PopupScreen "Tank 2S Status" 885x425
   TrendView "Trend view_1" at 280,6 size 600x360
   TextField "Text field_4" at 20,134 size 86x22; Text 'Pressure:'
   IOField "I/O field_1" at 175,129 size 90x25; FormatPattern s999.9; Unit  mBar
      ProcessValue <- "20_TANKS_IP_DATA_RIO_02_FIRST_TANK_TANKS_PRESS"
   TextField "Text field_5" at 20,168 size 113x22; Text 'Water Level:'
   IOField "I/O field_2" at 175,163 size 90x25; FormatPattern 999.9; Unit  %
      ProcessValue <- "20_TANKS_IP_DATA_RIO_02_SECOND_TANK_BWT_LEVEL"
   TextField "Text field_6" at 20,202 size 137x22; Text 'MBG Flow Rate:'
   IOField "I/O field_3" at 175,197 size 90x25; FormatPattern 999.9; Unit  m³/hr
      ProcessValue <- "20_TANKS_IP_DATA_RIO_02_SECOND_TANK_MBG_FLOW"
   TextField "Text field_7" at 20,236 size 135x22; Text 'USD Flow Rate:'
   IOField "I/O field_4" at 175,231 size 90x25; FormatPattern 999.9; Unit  m³/hr
      ProcessValue <- "20_TANKS_IP_DATA_RIO_02_SECOND_TANK_USD_FLOW"
   TextField "Text field_8" at 20,270 size 140x22; Text 'Water pH Level:'
   IOField "I/O field_5" at 175,265 size 90x25; FormatPattern 99.9
      ProcessValue <- "20_TANKS_IP_DATA_RIO_02_SECOND_TANK_BWT_PH"
   TextField "Text field_9" at 20,304 size 143x22; Text 'Water DO Level:'
   IOField "I/O field_6" at 175,299 size 90x25; FormatPattern 99.99; Unit  mg/l
      ProcessValue <- "20_TANKS_IP_DATA_RIO_02_SECOND_TANK_BWT_DO"
   TextField "Text field_10" at 20,338 size 174x22; Text 'Water Temperature:'
   IOField "I/O field_7" at 190,333 size 75x25; FormatPattern 999.9; Unit  °C
      ProcessValue <- "20_TANKS_IP_DATA_RIO_02_SECOND_TANK_BWT_TEMP"
   Button "Button_4" at 550,375 size 150x40; TextOff 'Disable Tank'; Authorization "Operate"
      on Press: function_b14e0dd5("504_Tank Grouping_DB2020_TANK ACTIV 5", 0)
   Button "Button_1" at 50,5 size 220x35; TextOff 'Starboard Tank 2 (2S)'
      on Release: function_efd93a16("Tank 2S Status", 168, 315, -1, 0, 1)
   TextField "Text field_1" at 20,90 size 109x25; Text 'TIME LEFT:'
   GraphicView "Graphic view_1" at 20,46 size 245x32; Picture "Tank Manually Disabled"
   GraphicIOField "Graphic I/O field_1" at 20,46 size 245x32; PictureList "Tank Process Stage_II"
      Visibility <- "504_Tank Grouping_DB2020_GROUP of TANK 5"
      ProcessValue <- "2110_BTCS_CNTRL_DB_BTCS_STATE"
   Button "Button_2" at 4,5 size 45x35; TextOff 'Text'; PictureOff "Graphic_286"
      on Click: function_efd93a16("Tank 2S Status", 0, 0, -1, -1, 1)
   Button "Button_3" at 287,375 size 230x40; TextOff 'Text'; Authorization "Operate"; PictureList "Water Level Override"
      on Press: InvertBit("2062_Warning_Data_Water Level Override 2S")
      ProcessValue <- "2062_Warning_Data_Water Level Override 2S"
   Button "Button_5" at 27,375 size 230x40; TextOff 'Tank Shutdown Alarm'
      Visibility <- "2062_Warning_Data_Alarm Tank S2"
   Button "Button_6" at 27,375 size 230x40; TextOff 'No/Low Water Level'; Authorization "Operate"
      Visibility <- "LT421 2S  TANK LEVEL ALARM_ALARM L"
   IOField "I/O field_29" at 218,90 size 47x25; FormatPattern 99; Unit m
      ProcessValue <- "504_Tank Grouping_DB2020_Time Left Tank_Time Left m Tank 5"
   IOField "I/O field_8" at 173,90 size 42x25; FormatPattern 99; Unit h
      ProcessValue <- "504_Tank Grouping_DB2020_Time Left Tank_Time Left h Tank 5"
   IOField "I/O field_9" at 128,90 size 42x25; FormatPattern 99; Unit d
      ProcessValue <- "504_Tank Grouping_DB2020_Time Left Tank_Time Left d Tank 5"

PopupScreen "Tank 3P Status" 885x425
   TrendView "Trend view_1" at 280,7 size 600x360
   TextField "Text field_4" at 20,135 size 86x22; Text 'Pressure:'
   IOField "I/O field_1" at 175,130 size 90x25; FormatPattern s999.9; Unit  mBar
      ProcessValue <- "20_TANKS_IP_DATA_RIO_03_FIRST_TANK_TANKS_PRESS"
   TextField "Text field_5" at 20,169 size 113x22; Text 'Water Level:'
   IOField "I/O field_2" at 175,164 size 90x25; FormatPattern 999.9; Unit  %
      ProcessValue <- "20_TANKS_IP_DATA_RIO_03_FIRST_TANK_BWT_LEVEL"
   TextField "Text field_6" at 20,203 size 137x22; Text 'MBG Flow Rate:'
   IOField "I/O field_3" at 175,198 size 90x25; FormatPattern 999.9; Unit  m³/hr
      ProcessValue <- "20_TANKS_IP_DATA_RIO_03_FIRST_TANK_MBG_FLOW"
   TextField "Text field_7" at 20,237 size 135x22; Text 'USD Flow Rate:'
   IOField "I/O field_4" at 175,232 size 90x25; FormatPattern 999.9; Unit  m³/hr
      ProcessValue <- "20_TANKS_IP_DATA_RIO_03_FIRST_TANK_USD_FLOW"
   TextField "Text field_8" at 20,271 size 140x22; Text 'Water pH Level:'
   IOField "I/O field_5" at 175,266 size 90x25; FormatPattern 99.9
      ProcessValue <- "20_TANKS_IP_DATA_RIO_03_FIRST_TANK_BWT_PH"
   TextField "Text field_9" at 20,305 size 143x22; Text 'Water DO Level:'
   IOField "I/O field_6" at 175,300 size 90x25; FormatPattern 99.99; Unit  mg/l
      ProcessValue <- "20_TANKS_IP_DATA_RIO_03_FIRST_TANK_BWT_DO"
   TextField "Text field_10" at 20,339 size 174x22; Text 'Water Temperature:'
   IOField "I/O field_7" at 190,334 size 75x25; FormatPattern 999.9; Unit  °C
      ProcessValue <- "20_TANKS_IP_DATA_RIO_03_FIRST_TANK_BWT_TEMP"
   Button "Button_4" at 545,375 size 150x40; TextOff 'Disable Tank'; Authorization "Operate"
      on Press: function_b14e0dd5("504_Tank Grouping_DB2020_TANK ACTIV 6", 0)
   Button "Button_1" at 51,5 size 220x35; TextOff 'Port Tank 3 (3P)'
      on Release: function_efd93a16("Tank 3P Status", 168, 315, -1, 0, 1)
   TextField "Text field_1" at 20,90 size 109x25; Text 'TIME LEFT:'
   GraphicView "Graphic view_1" at 20,46 size 245x32; Picture "Tank Manually Disabled"
   GraphicIOField "Graphic I/O field_1" at 20,46 size 245x32; PictureList "Tank Process Stage_II"
      Visibility <- "504_Tank Grouping_DB2020_GROUP of TANK 6"
      ProcessValue <- "2110_BTCS_CNTRL_DB_BTCS_STATE"
   Button "Button_2" at 4,5 size 45x35; TextOff 'Text'; PictureOff "Graphic_286"
      on Click: function_efd93a16("Tank 3P Status", 0, 0, -1, -1, 1)
   Button "Button_3" at 287,375 size 230x40; TextOff 'Text'; Authorization "Operate"; PictureList "Water Level Override"
      on Press: InvertBit("2062_Warning_Data_Water Level Override 3P")
      ProcessValue <- "2062_Warning_Data_Water Level Override 3P"
   Button "Button_5" at 27,375 size 230x40; TextOff 'Tank Shutdown Alarm'
      Visibility <- "2062_Warning_Data_Alarm Tank P3"
   Button "Button_6" at 27,375 size 230x40; TextOff 'No/Low Water Level'; Authorization "Operate"
      Visibility <- "LT422 3P  TANK LEVEL ALARM_ALARM L"
   IOField "I/O field_29" at 218,90 size 47x25; FormatPattern 99; Unit m
      ProcessValue <- "504_Tank Grouping_DB2020_Time Left Tank_Time Left m Tank 6"
   IOField "I/O field_8" at 173,90 size 42x25; FormatPattern 99; Unit h
      ProcessValue <- "504_Tank Grouping_DB2020_Time Left Tank_Time Left h Tank 6"
   IOField "I/O field_9" at 128,90 size 42x25; FormatPattern 99; Unit d
      ProcessValue <- "504_Tank Grouping_DB2020_Time Left Tank_Time Left d Tank 6"

PopupScreen "Tank 3S Status" 885x425
   TrendView "Trend view_1" at 280,7 size 600x360
   TextField "Text field_4" at 20,135 size 86x22; Text 'Pressure:'
   IOField "I/O field_1" at 175,130 size 90x25; FormatPattern s999.9; Unit  mBar
      ProcessValue <- "20_TANKS_IP_DATA_RIO_03_FIRST_TANK_TANKS_PRESS"
   TextField "Text field_5" at 20,169 size 113x22; Text 'Water Level:'
   IOField "I/O field_2" at 175,164 size 90x25; FormatPattern 999.9; Unit  %
      ProcessValue <- "20_TANKS_IP_DATA_RIO_03_SECOND_TANK_BWT_LEVEL"
   TextField "Text field_6" at 20,203 size 137x22; Text 'MBG Flow Rate:'
   IOField "I/O field_3" at 175,198 size 90x25; FormatPattern 999.9; Unit  m³/hr
      ProcessValue <- "20_TANKS_IP_DATA_RIO_03_SECOND_TANK_MBG_FLOW"
   TextField "Text field_7" at 20,237 size 135x22; Text 'USD Flow Rate:'
   IOField "I/O field_4" at 175,232 size 90x25; FormatPattern 999.9; Unit  m³/hr
      ProcessValue <- "20_TANKS_IP_DATA_RIO_03_SECOND_TANK_USD_FLOW"
   TextField "Text field_8" at 20,271 size 140x22; Text 'Water pH Level:'
   IOField "I/O field_5" at 175,266 size 90x25; FormatPattern 99.9
      ProcessValue <- "20_TANKS_IP_DATA_RIO_03_SECOND_TANK_BWT_PH"
   TextField "Text field_9" at 20,305 size 143x22; Text 'Water DO Level:'
   IOField "I/O field_6" at 175,300 size 90x25; FormatPattern 99.99; Unit  mg/l
      ProcessValue <- "20_TANKS_IP_DATA_RIO_03_SECOND_TANK_BWT_DO"
   TextField "Text field_10" at 20,339 size 174x22; Text 'Water Temperature:'
   IOField "I/O field_7" at 190,334 size 75x25; FormatPattern 999.9; Unit  °C
      ProcessValue <- "20_TANKS_IP_DATA_RIO_03_SECOND_TANK_BWT_TEMP"
   Button "Button_4" at 547,375 size 150x40; TextOff 'Disable Tank'; Authorization "Operate"
      on Press: function_b14e0dd5("504_Tank Grouping_DB2020_TANK ACTIV 7", 0)
   Button "Button_1" at 51,5 size 219x35; TextOff 'Starboard Tank 3 (3S)'
      on Release: function_efd93a16("Tank 3S Status", 168, 315, -1, 0, 1)
   TextField "Text field_1" at 20,90 size 109x25; Text 'TIME LEFT:'
   GraphicView "Graphic view_1" at 20,46 size 245x32; Picture "Tank Manually Disabled"
   GraphicIOField "Graphic I/O field_1" at 20,46 size 245x32; PictureList "Tank Process Stage_II"
      Visibility <- "504_Tank Grouping_DB2020_GROUP of TANK 7"
      ProcessValue <- "2110_BTCS_CNTRL_DB_BTCS_STATE"
   Button "Button_2" at 4,5 size 45x35; TextOff 'Text'; PictureOff "Graphic_286"
      on Click: function_efd93a16("Tank 3S Status", 0, 0, -1, -1, 1)
   Button "Button_3" at 287,375 size 230x40; TextOff 'Text'; Authorization "Operate"; PictureList "Water Level Override"
      on Press: InvertBit("2062_Warning_Data_Water Level Override 3S")
      ProcessValue <- "2062_Warning_Data_Water Level Override 3S"
   Button "Button_5" at 27,375 size 230x40; TextOff 'Tank Shutdown Alarm'
      Visibility <- "2062_Warning_Data_Alarm Tank S3"
   Button "Button_6" at 27,375 size 230x40; TextOff 'No/Low Water Level'; Authorization "Operate"
      Visibility <- "LT421 3S  TANK LEVEL ALARM_ALARM L"
   IOField "I/O field_29" at 218,90 size 47x25; FormatPattern 99; Unit m
      ProcessValue <- "504_Tank Grouping_DB2020_Time Left Tank_Time Left m Tank 7"
   IOField "I/O field_8" at 173,90 size 42x25; FormatPattern 99; Unit h
      ProcessValue <- "504_Tank Grouping_DB2020_Time Left Tank_Time Left h Tank 7"
   IOField "I/O field_9" at 128,90 size 42x25; FormatPattern 99; Unit d
      ProcessValue <- "504_Tank Grouping_DB2020_Time Left Tank_Time Left d Tank 7"

PopupScreen "Tank 4P Status" 885x425
   TrendView "Trend view_1" at 280,7 size 600x360
   TextField "Text field_4" at 20,135 size 86x22; Text 'Pressure:'
   IOField "I/O field_1" at 175,130 size 90x25; FormatPattern s999.9; Unit  mBar
      ProcessValue <- "20_TANKS_IP_DATA_RIO_04_FIRST_TANK_TANKS_PRESS"
   TextField "Text field_5" at 20,169 size 113x22; Text 'Water Level:'
   IOField "I/O field_2" at 175,164 size 90x25; FormatPattern 999.9; Unit  %
      ProcessValue <- "20_TANKS_IP_DATA_RIO_04_FIRST_TANK_BWT_LEVEL"
   TextField "Text field_6" at 20,203 size 137x22; Text 'MBG Flow Rate:'
   IOField "I/O field_3" at 175,198 size 90x25; FormatPattern 999.9; Unit  m³/hr
      ProcessValue <- "20_TANKS_IP_DATA_RIO_04_FIRST_TANK_MBG_FLOW"
   TextField "Text field_7" at 20,237 size 135x22; Text 'USD Flow Rate:'
   IOField "I/O field_4" at 175,232 size 90x25; FormatPattern 999.9; Unit  m³/hr
      ProcessValue <- "20_TANKS_IP_DATA_RIO_04_FIRST_TANK_USD_FLOW"
   TextField "Text field_8" at 20,271 size 140x22; Text 'Water pH Level:'
   IOField "I/O field_5" at 175,266 size 90x25; FormatPattern 99.9
      ProcessValue <- "20_TANKS_IP_DATA_RIO_04_FIRST_TANK_BWT_PH"
   TextField "Text field_9" at 20,305 size 143x22; Text 'Water DO Level:'
   IOField "I/O field_6" at 175,300 size 90x25; FormatPattern 99.99; Unit  mg/l
      ProcessValue <- "20_TANKS_IP_DATA_RIO_04_FIRST_TANK_BWT_DO"
   TextField "Text field_10" at 20,339 size 174x22; Text 'Water Temperature:'
   IOField "I/O field_7" at 190,334 size 75x25; FormatPattern 999.9; Unit  °C
      ProcessValue <- "20_TANKS_IP_DATA_RIO_04_FIRST_TANK_BWT_TEMP"
   Button "Button_4" at 545,375 size 150x40; TextOff 'Disable Tank'; Authorization "Operate"
      on Press: function_b14e0dd5("504_Tank Grouping_DB2020_TANK ACTIV 8", 0)
   Button "Button_1" at 51,5 size 219x35; TextOff 'Port Tank 4 (4P)'
      on Release: function_efd93a16("Tank 4P Status", 168, 315, -1, 2, 1)
   TextField "Text field_1" at 20,90 size 109x25; Text 'TIME LEFT:'
   GraphicView "Graphic view_1" at 20,46 size 245x32; Picture "Tank Manually Disabled"
   GraphicIOField "Graphic I/O field_1" at 20,46 size 245x32; PictureList "Tank Process Stage_II"
      Visibility <- "504_Tank Grouping_DB2020_GROUP of TANK 8"
      ProcessValue <- "2110_BTCS_CNTRL_DB_BTCS_STATE"
   Button "Button_2" at 4,5 size 45x35; TextOff 'Text'; PictureOff "Graphic_286"
      on Click: function_efd93a16("Tank 4P Status", 0, 0, -1, -1, 1)
   Button "Button_3" at 287,375 size 230x40; TextOff 'Text'; Authorization "Operate"; PictureList "Water Level Override"
      on Press: InvertBit("2062_Warning_Data_Water Level Override 4P")
      ProcessValue <- "2062_Warning_Data_Water Level Override 4P"
   Button "Button_5" at 27,375 size 230x40; TextOff 'Tank Shutdown Alarm'
      Visibility <- "2062_Warning_Data_Alarm Tank P4"
   Button "Button_6" at 27,375 size 230x40; TextOff 'No/Low Water Level'; Authorization "Operate"
      Visibility <- "LT422 4P  TANK LEVEL ALARM_ALARM L"
   IOField "I/O field_29" at 218,90 size 47x25; FormatPattern 99; Unit m
      ProcessValue <- "504_Tank Grouping_DB2020_Time Left Tank_Time Left m Tank 8"
   IOField "I/O field_8" at 173,90 size 42x25; FormatPattern 99; Unit h
      ProcessValue <- "504_Tank Grouping_DB2020_Time Left Tank_Time Left h Tank 8"
   IOField "I/O field_9" at 128,90 size 42x25; FormatPattern 99; Unit d
      ProcessValue <- "504_Tank Grouping_DB2020_Time Left Tank_Time Left d Tank 8"

PopupScreen "Tank 4S Status" 885x425
   TrendView "Trend view_1" at 280,7 size 600x360
   TextField "Text field_4" at 20,135 size 86x22; Text 'Pressure:'
   IOField "I/O field_1" at 175,130 size 90x25; FormatPattern s999.9; Unit  mBar
      ProcessValue <- "20_TANKS_IP_DATA_RIO_04_FIRST_TANK_TANKS_PRESS"
   TextField "Text field_5" at 20,169 size 113x22; Text 'Water Level:'
   IOField "I/O field_2" at 175,164 size 90x25; FormatPattern 999.9; Unit  %
      ProcessValue <- "20_TANKS_IP_DATA_RIO_04_SECOND_TANK_BWT_LEVEL"
   TextField "Text field_6" at 20,203 size 137x22; Text 'MBG Flow Rate:'
   IOField "I/O field_3" at 175,198 size 90x25; FormatPattern 999.9; Unit  m³/hr
      ProcessValue <- "20_TANKS_IP_DATA_RIO_04_SECOND_TANK_MBG_FLOW"
   TextField "Text field_7" at 20,237 size 135x22; Text 'USD Flow Rate:'
   IOField "I/O field_4" at 175,232 size 90x25; FormatPattern 999.9; Unit  m³/hr
      ProcessValue <- "20_TANKS_IP_DATA_RIO_04_SECOND_TANK_USD_FLOW"
   TextField "Text field_8" at 20,271 size 140x22; Text 'Water pH Level:'
   IOField "I/O field_5" at 175,266 size 90x25; FormatPattern 99.9
      ProcessValue <- "20_TANKS_IP_DATA_RIO_04_SECOND_TANK_BWT_PH"
   TextField "Text field_9" at 20,305 size 143x22; Text 'Water DO Level:'
   IOField "I/O field_6" at 175,300 size 90x25; FormatPattern 99.99; Unit  mg/l
      ProcessValue <- "20_TANKS_IP_DATA_RIO_04_SECOND_TANK_BWT_DO"
   TextField "Text field_10" at 20,339 size 174x22; Text 'Water Temperature:'
   IOField "I/O field_7" at 190,334 size 75x25; FormatPattern 999.9; Unit  °C
      ProcessValue <- "20_TANKS_IP_DATA_RIO_04_SECOND_TANK_BWT_TEMP"
   Button "Button_4" at 545,375 size 150x40; TextOff 'Disable Tank'; Authorization "Operate"
      on Press: function_b14e0dd5("504_Tank Grouping_DB2020_TANK ACTIV 9", 0)
   Button "Button_1" at 50,5 size 220x35; TextOff 'Starboard Tank 4 (4S)'
      on Release: function_efd93a16("Tank 4S Status", 168, 315, -1, 2, 1)
   TextField "Text field_1" at 20,90 size 109x25; Text 'TIME LEFT:'
   GraphicView "Graphic view_1" at 20,46 size 245x32; Picture "Tank Manually Disabled"
   GraphicIOField "Graphic I/O field_1" at 20,46 size 245x32; PictureList "Tank Process Stage_II"
      Visibility <- "504_Tank Grouping_DB2020_GROUP of TANK 9"
      ProcessValue <- "2110_BTCS_CNTRL_DB_BTCS_STATE"
   Button "Button_2" at 4,5 size 45x35; TextOff 'Text'; PictureOff "Graphic_286"
      on Click: function_efd93a16("Tank 4S Status", 0, 0, -1, -1, 1)
   Button "Button_3" at 287,375 size 230x40; TextOff 'Text'; Authorization "Operate"; PictureList "Water Level Override"
      on Press: InvertBit("2062_Warning_Data_Water Level Override 4S")
      ProcessValue <- "2062_Warning_Data_Water Level Override 4S"
   Button "Button_5" at 27,375 size 230x40; TextOff 'Tank Shutdown Alarm'
      Visibility <- "2062_Warning_Data_Alarm Tank S4"
   Button "Button_6" at 27,375 size 230x40; TextOff 'No/Low Water Level'; Authorization "Operate"
      Visibility <- "LT421 4S  TANK LEVEL ALARM_ALARM L"
   IOField "I/O field_29" at 218,90 size 47x25; FormatPattern 99; Unit m
      ProcessValue <- "504_Tank Grouping_DB2020_Time Left Tank_Time Left m Tank 9"
   IOField "I/O field_8" at 173,90 size 42x25; FormatPattern 99; Unit h
      ProcessValue <- "504_Tank Grouping_DB2020_Time Left Tank_Time Left h Tank 9"
   IOField "I/O field_9" at 128,90 size 42x25; FormatPattern 99; Unit d
      ProcessValue <- "504_Tank Grouping_DB2020_Time Left Tank_Time Left d Tank 9"

PopupScreen "Tank 5P Status" 885x425
   TrendView "Trend view_1" at 280,7 size 600x360
   TextField "Text field_4" at 20,135 size 86x22; Text 'Pressure:'
   IOField "I/O field_1" at 175,130 size 90x25; FormatPattern s999.9; Unit  mBar
      ProcessValue <- "20_TANKS_IP_DATA_RIO_05_FIRST_TANK_TANKS_PRESS"
   TextField "Text field_5" at 20,169 size 113x22; Text 'Water Level:'
   IOField "I/O field_2" at 175,164 size 90x25; FormatPattern 999.9; Unit  %
      ProcessValue <- "20_TANKS_IP_DATA_RIO_05_FIRST_TANK_BWT_LEVEL"
   TextField "Text field_6" at 20,203 size 137x22; Text 'MBG Flow Rate:'
   IOField "I/O field_3" at 175,198 size 90x25; FormatPattern 999.9; Unit  m³/hr
      ProcessValue <- "20_TANKS_IP_DATA_RIO_05_FIRST_TANK_MBG_FLOW"
   TextField "Text field_7" at 20,237 size 135x22; Text 'USD Flow Rate:'
   IOField "I/O field_4" at 175,232 size 90x25; FormatPattern 999.9; Unit  m³/hr
      ProcessValue <- "20_TANKS_IP_DATA_RIO_05_FIRST_TANK_USD_FLOW"
   TextField "Text field_8" at 20,271 size 140x22; Text 'Water pH Level:'
   IOField "I/O field_5" at 175,266 size 90x25; FormatPattern 99.9
      ProcessValue <- "20_TANKS_IP_DATA_RIO_05_FIRST_TANK_BWT_PH"
   TextField "Text field_9" at 20,305 size 143x22; Text 'Water DO Level:'
   IOField "I/O field_6" at 175,300 size 90x25; FormatPattern 99.99; Unit  mg/l
      ProcessValue <- "20_TANKS_IP_DATA_RIO_05_FIRST_TANK_BWT_DO"
   TextField "Text field_10" at 20,339 size 174x22; Text 'Water Temperature:'
   IOField "I/O field_7" at 190,334 size 75x25; FormatPattern 999.9; Unit  °C
      ProcessValue <- "20_TANKS_IP_DATA_RIO_05_FIRST_TANK_BWT_TEMP"
   Button "Button_4" at 546,375 size 150x40; TextOff 'Disable Tank'; Authorization "Operate"
      on Press: function_b14e0dd5("504_Tank Grouping_DB2020_TANK ACTIV 10", 0)
   Button "Button_1" at 51,5 size 219x35; TextOff 'Port Tank 5 (5P)'
      on Release: function_efd93a16("Tank 5P Status", 168, 315, -1, 2, 1)
   TextField "Text field_1" at 20,90 size 109x25; Text 'TIME LEFT:'
   GraphicView "Graphic view_1" at 20,46 size 245x32; Picture "Tank Manually Disabled"
   GraphicIOField "Graphic I/O field_1" at 20,46 size 245x32; PictureList "Tank Process Stage_II"
      Visibility <- "504_Tank Grouping_DB2020_GROUP of TANK 10"
      ProcessValue <- "2110_BTCS_CNTRL_DB_BTCS_STATE"
   Button "Button_2" at 4,5 size 45x35; TextOff 'Text'; PictureOff "Graphic_286"
      on Click: function_efd93a16("Tank 5P Status", 0, 0, -1, -1, 1)
   Button "Button_3" at 287,375 size 230x40; TextOff 'Text'; Authorization "Operate"; PictureList "Water Level Override"
      on Press: InvertBit("2062_Warning_Data_Water Level Override 5P")
      ProcessValue <- "2062_Warning_Data_Water Level Override 5P"
   Button "Button_5" at 27,375 size 230x40; TextOff 'Tank Shutdown Alarm'
      Visibility <- "2062_Warning_Data_Alarm Tank P5"
   Button "Button_6" at 27,375 size 230x40; TextOff 'No/Low Water Level'; Authorization "Operate"
      Visibility <- "LT422 5P  TANK LEVEL ALARM_ALARM L"
   IOField "I/O field_29" at 218,90 size 47x25; FormatPattern 99; Unit m
      ProcessValue <- "504_Tank Grouping_DB2020_Time Left Tank_Time Left m Tank 10"
   IOField "I/O field_8" at 173,90 size 42x25; FormatPattern 99; Unit h
      ProcessValue <- "504_Tank Grouping_DB2020_Time Left Tank_Time Left h Tank 10"
   IOField "I/O field_9" at 128,90 size 42x25; FormatPattern 99; Unit d
      ProcessValue <- "504_Tank Grouping_DB2020_Time Left Tank_Time Left d Tank 10"

PopupScreen "Tank 5S Status" 885x425
   TrendView "Trend view_1" at 280,7 size 600x360
   TextField "Text field_4" at 20,135 size 86x22; Text 'Pressure:'
   IOField "I/O field_1" at 175,130 size 90x25; FormatPattern s999.9; Unit  mBar
      ProcessValue <- "20_TANKS_IP_DATA_RIO_05_FIRST_TANK_TANKS_PRESS"
   TextField "Text field_5" at 20,169 size 113x22; Text 'Water Level:'
   IOField "I/O field_2" at 175,164 size 90x25; FormatPattern 999.9; Unit  %
      ProcessValue <- "20_TANKS_IP_DATA_RIO_05_SECOND_TANK_BWT_LEVEL"
   TextField "Text field_6" at 20,203 size 137x22; Text 'MBG Flow Rate:'
   IOField "I/O field_3" at 175,198 size 90x25; FormatPattern 999.9; Unit  m³/hr
      ProcessValue <- "20_TANKS_IP_DATA_RIO_05_SECOND_TANK_MBG_FLOW"
   TextField "Text field_7" at 20,237 size 135x22; Text 'USD Flow Rate:'
   IOField "I/O field_4" at 175,232 size 90x25; FormatPattern 999.9; Unit  m³/hr
      ProcessValue <- "20_TANKS_IP_DATA_RIO_05_SECOND_TANK_USD_FLOW"
   TextField "Text field_8" at 20,271 size 140x22; Text 'Water pH Level:'
   IOField "I/O field_5" at 175,266 size 90x25; FormatPattern 99.9
      ProcessValue <- "20_TANKS_IP_DATA_RIO_05_SECOND_TANK_BWT_PH"
   TextField "Text field_9" at 20,305 size 143x22; Text 'Water DO Level:'
   IOField "I/O field_6" at 175,300 size 90x25; FormatPattern 99.99; Unit  mg/l
      ProcessValue <- "20_TANKS_IP_DATA_RIO_05_SECOND_TANK_BWT_DO"
   TextField "Text field_10" at 20,339 size 174x22; Text 'Water Temperature:'
   IOField "I/O field_7" at 190,334 size 75x25; FormatPattern 999.9; Unit  °C
      ProcessValue <- "20_TANKS_IP_DATA_RIO_05_SECOND_TANK_BWT_TEMP"
   Button "Button_4" at 550,375 size 150x40; TextOff 'Disable Tank'; Authorization "Operate"
      on Press: function_b14e0dd5("504_Tank Grouping_DB2020_TANK ACTIV 11", 0)
   Button "Button_1" at 50,5 size 220x35; TextOff 'Starboard Tank 5 (5S)'
      on Release: function_efd93a16("Tank 5S Status", 168, 315, -1, 2, 1)
   TextField "Text field_1" at 20,90 size 109x25; Text 'TIME LEFT:'
   GraphicView "Graphic view_1" at 20,46 size 245x32; Picture "Tank Manually Disabled"
   GraphicIOField "Graphic I/O field_1" at 20,46 size 245x32; PictureList "Tank Process Stage_II"
      Visibility <- "504_Tank Grouping_DB2020_GROUP of TANK 11"
      ProcessValue <- "2110_BTCS_CNTRL_DB_BTCS_STATE"
   Button "Button_2" at 4,5 size 45x35; TextOff 'Text'; PictureOff "Graphic_286"
      on Click: function_efd93a16("Tank 5S Status", 0, 0, -1, -1, 1)
   Button "Button_3" at 287,375 size 230x40; TextOff 'Text'; Authorization "Operate"; PictureList "Water Level Override"
      on Press: InvertBit("2062_Warning_Data_Water Level Override 5S")
      ProcessValue <- "2062_Warning_Data_Water Level Override 5S"
   Button "Button_5" at 27,375 size 230x40; TextOff 'Tank Shutdown Alarm'
      Visibility <- "2062_Warning_Data_Alarm Tank S5"
   Button "Button_6" at 27,375 size 230x40; TextOff 'No/Low Water Level'; Authorization "Operate"
      Visibility <- "LT421 5S  TANK LEVEL ALARM_ALARM L"
   IOField "I/O field_29" at 218,90 size 47x25; FormatPattern 99; Unit m
      ProcessValue <- "504_Tank Grouping_DB2020_Time Left Tank_Time Left m Tank 11"
   IOField "I/O field_8" at 173,90 size 42x25; FormatPattern 99; Unit h
      ProcessValue <- "504_Tank Grouping_DB2020_Time Left Tank_Time Left h Tank 11"
   IOField "I/O field_9" at 128,90 size 42x25; FormatPattern 99; Unit d
      ProcessValue <- "504_Tank Grouping_DB2020_Time Left Tank_Time Left d Tank 11"

PopupScreen "Tank 6P Status" 885x425
   TrendView "Trend view_1" at 280,7 size 600x360
   TextField "Text field_4" at 20,135 size 86x22; Text 'Pressure:'
   IOField "I/O field_1" at 175,130 size 90x25; FormatPattern s999.9; Unit  mBar
      ProcessValue <- "20_TANKS_IP_DATA_RIO_06_FIRST_TANK_TANKS_PRESS"
   TextField "Text field_5" at 20,169 size 113x22; Text 'Water Level:'
   IOField "I/O field_2" at 175,164 size 90x25; FormatPattern 999.9; Unit  %
      ProcessValue <- "20_TANKS_IP_DATA_RIO_06_FIRST_TANK_BWT_LEVEL"
   TextField "Text field_6" at 20,203 size 137x22; Text 'MBG Flow Rate:'
   IOField "I/O field_3" at 175,198 size 90x25; FormatPattern 999.9; Unit  m³/hr
      ProcessValue <- "20_TANKS_IP_DATA_RIO_06_FIRST_TANK_MBG_FLOW"
   TextField "Text field_7" at 20,237 size 135x22; Text 'USD Flow Rate:'
   IOField "I/O field_4" at 175,232 size 90x25; FormatPattern 999.9; Unit  m³/hr
      ProcessValue <- "20_TANKS_IP_DATA_RIO_06_FIRST_TANK_USD_FLOW"
   TextField "Text field_8" at 20,271 size 140x22; Text 'Water pH Level:'
   IOField "I/O field_5" at 175,266 size 90x25; FormatPattern 99.9
      ProcessValue <- "20_TANKS_IP_DATA_RIO_06_FIRST_TANK_BWT_PH"
   TextField "Text field_9" at 20,305 size 143x22; Text 'Water DO Level:'
   IOField "I/O field_6" at 175,300 size 90x25; FormatPattern 99.99; Unit  mg/l
      ProcessValue <- "20_TANKS_IP_DATA_RIO_06_FIRST_TANK_BWT_DO"
   TextField "Text field_10" at 20,339 size 174x22; Text 'Water Temperature:'
   IOField "I/O field_7" at 190,334 size 75x25; FormatPattern 999.9; Unit  °C
      ProcessValue <- "20_TANKS_IP_DATA_RIO_06_FIRST_TANK_BWT_TEMP"
   Button "Button_4" at 542,374 size 150x40; TextOff 'Disable Tank'; Authorization "Operate"
      on Press: function_b14e0dd5("504_Tank Grouping_DB2020_TANK ACTIV 12", 0)
   Button "Button_1" at 51,5 size 219x35; TextOff 'Port Tank 6 (6P)'
      on Release: function_efd93a16("Tank 6P Status", 168, 315, -1, 2, 1)
   TextField "Text field_1" at 20,90 size 109x25; Text 'TIME LEFT:'
   GraphicView "Graphic view_1" at 20,46 size 245x32; Picture "Tank Manually Disabled"
   GraphicIOField "Graphic I/O field_1" at 20,46 size 245x32; PictureList "Tank Process Stage_II"
      Visibility <- "504_Tank Grouping_DB2020_GROUP of TANK 12"
      ProcessValue <- "2110_BTCS_CNTRL_DB_BTCS_STATE"
   Button "Button_2" at 4,5 size 45x35; TextOff 'Text'; PictureOff "Graphic_286"
      on Click: function_efd93a16("Tank 6P Status", 0, 0, -1, -1, 1)
   Button "Button_3" at 287,375 size 230x40; TextOff 'Text'; Authorization "Operate"; PictureList "Water Level Override"
      on Press: InvertBit("2062_Warning_Data_Water Level Override 6P")
      ProcessValue <- "2062_Warning_Data_Water Level Override 6P"
   Button "Button_5" at 27,375 size 230x40; TextOff 'Tank Shutdown Alarm'
      Visibility <- "2062_Warning_Data_Alarm Tank P6"
   Button "Button_6" at 27,375 size 230x40; TextOff 'No/Low Water Level'; Authorization "Operate"
      Visibility <- "LT422 6P  TANK LEVEL ALARM_ALARM L"
   IOField "I/O field_29" at 218,90 size 47x25; FormatPattern 99; Unit m
      ProcessValue <- "504_Tank Grouping_DB2020_Time Left Tank_Time Left m Tank 12"
   IOField "I/O field_8" at 173,90 size 42x25; FormatPattern 99; Unit h
      ProcessValue <- "504_Tank Grouping_DB2020_Time Left Tank_Time Left h Tank 12"
   IOField "I/O field_9" at 128,90 size 42x25; FormatPattern 99; Unit d
      ProcessValue <- "504_Tank Grouping_DB2020_Time Left Tank_Time Left d Tank 12"

PopupScreen "Tank 6S Status" 885x425
   TrendView "Trend view_1" at 280,7 size 600x360
   TextField "Text field_4" at 20,135 size 86x22; Text 'Pressure:'
   IOField "I/O field_1" at 175,130 size 90x25; FormatPattern s999.9; Unit  mBar
      ProcessValue <- "20_TANKS_IP_DATA_RIO_06_FIRST_TANK_TANKS_PRESS"
   TextField "Text field_5" at 20,169 size 113x22; Text 'Water Level:'
   IOField "I/O field_2" at 175,164 size 90x25; FormatPattern 999.9; Unit  %
      ProcessValue <- "20_TANKS_IP_DATA_RIO_06_SECOND_TANK_BWT_LEVEL"
   TextField "Text field_6" at 20,203 size 137x22; Text 'MBG Flow Rate:'
   IOField "I/O field_3" at 175,198 size 90x25; FormatPattern 999.9; Unit  m³/hr
      ProcessValue <- "20_TANKS_IP_DATA_RIO_06_SECOND_TANK_MBG_FLOW"
   TextField "Text field_7" at 20,237 size 135x22; Text 'USD Flow Rate:'
   IOField "I/O field_4" at 175,232 size 90x25; FormatPattern 999.9; Unit  m³/hr
      ProcessValue <- "20_TANKS_IP_DATA_RIO_06_SECOND_TANK_USD_FLOW"
   TextField "Text field_8" at 20,271 size 140x22; Text 'Water pH Level:'
   IOField "I/O field_5" at 175,266 size 90x25; FormatPattern 99.9
      ProcessValue <- "20_TANKS_IP_DATA_RIO_06_SECOND_TANK_BWT_PH"
   TextField "Text field_9" at 20,305 size 143x22; Text 'Water DO Level:'
   IOField "I/O field_6" at 175,300 size 90x25; FormatPattern 99.99; Unit  mg/l
      ProcessValue <- "20_TANKS_IP_DATA_RIO_06_SECOND_TANK_BWT_DO"
   TextField "Text field_10" at 20,339 size 174x22; Text 'Water Temperature:'
   IOField "I/O field_7" at 190,334 size 75x25; FormatPattern 999.9; Unit  °C
      ProcessValue <- "20_TANKS_IP_DATA_RIO_06_SECOND_TANK_BWT_TEMP"
   Button "Button_4" at 545,377 size 150x40; TextOff 'Disable Tank'; Authorization "Operate"
      on Press: function_b14e0dd5("504_Tank Grouping_DB2020_TANK ACTIV 13", 0)
   Button "Button_1" at 51,5 size 219x35; TextOff 'Starboard Tank 6 (6S)'
      on Release: function_efd93a16("Tank 6S Status", 168, 315, -1, 2, 1)
   TextField "Text field_1" at 20,90 size 109x25; Text 'TIME LEFT:'
   GraphicView "Graphic view_1" at 20,46 size 245x32; Picture "Tank Manually Disabled"
   GraphicIOField "Graphic I/O field_1" at 20,46 size 245x32; PictureList "Tank Process Stage_II"
      Visibility <- "504_Tank Grouping_DB2020_GROUP of TANK 13"
      ProcessValue <- "2110_BTCS_CNTRL_DB_BTCS_STATE"
   Button "Button_2" at 4,5 size 45x35; TextOff 'Text'; PictureOff "Graphic_286"
      on Click: function_efd93a16("Tank 6S Status", 0, 0, -1, -1, 1)
   Button "Button_3" at 287,375 size 230x40; TextOff 'Text'; Authorization "Operate"; PictureList "Water Level Override"
      on Press: InvertBit("2062_Warning_Data_Water Level Override 6S")
      ProcessValue <- "2062_Warning_Data_Water Level Override 6S"
   Button "Button_5" at 27,375 size 230x40; TextOff 'Tank Shutdown Alarm'
      Visibility <- "2062_Warning_Data_Alarm Tank S6"
   Button "Button_6" at 27,375 size 230x40; TextOff 'No/Low Water Level'; Authorization "Operate"
      Visibility <- "LT421 6S  TANK LEVEL ALARM_ALARM L"
   IOField "I/O field_29" at 218,90 size 47x25; FormatPattern 99; Unit m
      ProcessValue <- "504_Tank Grouping_DB2020_Time Left Tank_Time Left m Tank 13"
   IOField "I/O field_8" at 173,90 size 42x25; FormatPattern 99; Unit h
      ProcessValue <- "504_Tank Grouping_DB2020_Time Left Tank_Time Left h Tank 13"
   IOField "I/O field_9" at 128,90 size 42x25; FormatPattern 99; Unit d
      ProcessValue <- "504_Tank Grouping_DB2020_Time Left Tank_Time Left d Tank 13"

PopupScreen "Tank AP Status" 885x425
   TrendView "Trend view_1" at 280,7 size 600x360
   TextField "Text field_4" at 20,135 size 86x22; Text 'Pressure:'
   IOField "I/O field_1" at 175,130 size 90x25; FormatPattern s999.9; Unit  mBar
      ProcessValue <- "20_TANKS_IP_DATA_RIO_07_FIRST_TANK_TANKS_PRESS"
   TextField "Text field_5" at 20,169 size 113x22; Text 'Water Level:'
   IOField "I/O field_2" at 175,164 size 90x25; FormatPattern 999.9; Unit  %
      ProcessValue <- "20_TANKS_IP_DATA_RIO_07_FIRST_TANK_BWT_LEVEL"
   TextField "Text field_6" at 20,203 size 137x22; Text 'MBG Flow Rate:'
   IOField "I/O field_3" at 175,198 size 90x25; FormatPattern 999.9; Unit  m³/hr
      ProcessValue <- "20_TANKS_IP_DATA_RIO_07_FIRST_TANK_MBG_FLOW"
   TextField "Text field_7" at 20,237 size 135x22; Text 'USD Flow Rate:'
   IOField "I/O field_4" at 175,232 size 90x25; FormatPattern 999.9; Unit  m³/hr
      ProcessValue <- "20_TANKS_IP_DATA_RIO_07_FIRST_TANK_USD_FLOW"
   TextField "Text field_8" at 20,271 size 140x22; Text 'Water pH Level:'
   IOField "I/O field_5" at 175,266 size 90x25; FormatPattern 99.9
      ProcessValue <- "20_TANKS_IP_DATA_RIO_07_FIRST_TANK_BWT_PH"
   TextField "Text field_9" at 20,305 size 143x22; Text 'Water DO Level:'
   IOField "I/O field_6" at 175,300 size 90x25; FormatPattern 99.99; Unit  mg/l
      ProcessValue <- "20_TANKS_IP_DATA_RIO_07_FIRST_TANK_BWT_DO"
   TextField "Text field_10" at 20,339 size 174x22; Text 'Water Temperature:'
   IOField "I/O field_7" at 190,334 size 75x25; FormatPattern 999.9; Unit  °C
      ProcessValue <- "20_TANKS_IP_DATA_RIO_07_FIRST_TANK_BWT_TEMP"
   Button "Button_4" at 538,375 size 150x40; TextOff 'Disable Tank'; Authorization "Operate"
      on Press: function_b14e0dd5("504_Tank Grouping_DB2020_TANK ACTIV 14", 0)
   Button "Button_1" at 51,5 size 219x35; TextOff 'Aft Peak Tank (APT)'
      on Release: function_efd93a16("Tank AP Status", 168, 315, -1, 2, 1)
   TextField "Text field_1" at 20,90 size 109x25; Text 'TIME LEFT:'
   GraphicView "Graphic view_1" at 20,46 size 245x32; Picture "Tank Manually Disabled"
   GraphicIOField "Graphic I/O field_1" at 20,46 size 245x32; PictureList "Tank Process Stage_II"
      Visibility <- "504_Tank Grouping_DB2020_GROUP of TANK 14"
      ProcessValue <- "2110_BTCS_CNTRL_DB_BTCS_STATE"
   Button "Button_2" at 4,5 size 45x35; TextOff 'Text'; PictureOff "Graphic_286"
      on Click: function_efd93a16("Tank AP Status", 0, 0, -1, -1, 1)
   Button "Button_3" at 287,375 size 230x40; TextOff 'Text'; Authorization "Operate"; PictureList "Water Level Override"
      on Press: InvertBit("2062_Warning_Data_Water Level Override APT")
      ProcessValue <- "2062_Warning_Data_Water Level Override APT"
   Button "Button_5" at 27,375 size 230x40; TextOff 'Tank Shutdown Alarm'
      Visibility <- "2062_Warning_Data_Alarm Tank APT"
   Button "Button_6" at 27,375 size 230x40; TextOff 'No/Low Water Level'; Authorization "Operate"
      Visibility <- "LT422 APT  TANK LEVEL ALARM_ALARM L"
   IOField "I/O field_29" at 218,90 size 47x25; FormatPattern 99; Unit m
      ProcessValue <- "504_Tank Grouping_DB2020_Time Left Tank_Time Left m Tank 14"
   IOField "I/O field_8" at 173,90 size 42x25; FormatPattern 99; Unit h
      ProcessValue <- "504_Tank Grouping_DB2020_Time Left Tank_Time Left h Tank 14"
   IOField "I/O field_9" at 128,90 size 42x25; FormatPattern 99; Unit d
      ProcessValue <- "504_Tank Grouping_DB2020_Time Left Tank_Time Left d Tank 14"

PopupScreen "Tank FP Status" 885x425
   TrendView "Trend view_1" at 280,7 size 600x360
   TextField "Text field_1" at 20,90 size 109x25; Text 'TIME LEFT:'
   TextField "Text field_4" at 20,135 size 86x22; Text 'Pressure:'
   IOField "I/O field_1" at 175,130 size 90x25; FormatPattern s999.9; Unit  mBar
      ProcessValue <- "20_TANKS_IP_DATA_RIO_01_FIRST_TANK_TANKS_PRESS"
   TextField "Text field_5" at 20,169 size 113x22; Text 'Water Level:'
   IOField "I/O field_2" at 175,164 size 90x25; FormatPattern 999.9; Unit  %
      ProcessValue <- "20_TANKS_IP_DATA_RIO_01_FIRST_TANK_BWT_LEVEL"
   TextField "Text field_6" at 20,203 size 137x22; Text 'MBG Flow Rate:'
   IOField "I/O field_3" at 175,198 size 90x25; FormatPattern 999.9; Unit  m³/hr
      ProcessValue <- "20_TANKS_IP_DATA_RIO_01_FIRST_TANK_MBG_FLOW"
   TextField "Text field_7" at 20,237 size 135x22; Text 'USD Flow Rate:'
   IOField "I/O field_4" at 175,232 size 90x25; FormatPattern 999.9; Unit  m³/hr
      ProcessValue <- "20_TANKS_IP_DATA_RIO_01_FIRST_TANK_USD_FLOW"
   TextField "Text field_8" at 20,271 size 140x22; Text 'Water pH Level:'
   IOField "I/O field_5" at 175,266 size 90x25; FormatPattern 99.9
      ProcessValue <- "20_TANKS_IP_DATA_RIO_01_FIRST_TANK_BWT_PH"
   TextField "Text field_9" at 20,305 size 143x22; Text 'Water DO Level:'
   IOField "I/O field_6" at 175,300 size 90x25; FormatPattern 99.99; Unit  mg/l
      ProcessValue <- "20_TANKS_IP_DATA_RIO_01_FIRST_TANK_BWT_DO"
   TextField "Text field_10" at 20,339 size 174x22; Text 'Water Temperature:'
   IOField "I/O field_7" at 190,334 size 75x25; FormatPattern 999.9; Unit  °C
      ProcessValue <- "20_TANKS_IP_DATA_RIO_01_FIRST_TANK_BWT_TEMP"
   IOField "I/O field_29" at 218,90 size 47x25; FormatPattern 99; Unit m
      ProcessValue <- "504_Tank Grouping_DB2020_Time Left Tank_Time Left m Tank 1"
   Button "Button_2" at 712,375 size 150x40; TextOff 'Reset Tank'
      Visibility <- "AlwaysTRUE"
   Button "Button_3" at 287,375 size 230x40; TextOff 'Text'; Authorization "Operate"; PictureList "Water Level Override"
      on Press: InvertBit("2062_Warning_Data_Water Level Override FPT")
      ProcessValue <- "2062_Warning_Data_Water Level Override FPT"
   Button "Button_4" at 539,375 size 150x40; TextOff 'Disable Tank'; Authorization "Operate"
      on Press: function_b14e0dd5("504_Tank Grouping_DB2020_TANK ACTIV 1", 0)
   Button "Button_5" at 27,375 size 230x40; TextOff 'Tank Shutdown Alarm'
      ProcessValue <- "2062_Warning_Data_Water Level Override FPT"
      Visibility <- "2062_Warning_Data_Alarm Tank FPT"
   Button "Button_6" at 27,375 size 230x40; TextOff 'No/Low Water Level'
      ProcessValue <- "2062_Warning_Data_Water Level Override FPT"
      Visibility <- "LT422 FPT  TANK LEVEL ALARM_ALARM L"
   GraphicView "Graphic view_1" at 20,46 size 245x32; Picture "Tank Manually Disabled"
   Button "Button_1" at 51,5 size 219x35; TextOff 'Fore Peak Tank (FPT)'
   GraphicIOField "Graphic I/O field_1" at 20,46 size 245x32; PictureList "Tank Process Stage_II"
      Visibility <- "504_Tank Grouping_DB2020_GROUP of TANK 1"
      ProcessValue <- "2110_BTCS_CNTRL_DB_BTCS_STATE"
   Button "Button_7" at 4,5 size 45x35; TextOff 'Text'; PictureOff "Graphic_286"
      on Click: function_efd93a16("Tank FP Status", 0, 0, -1, -1, 1)
   IOField "I/O field_8" at 173,90 size 42x25; FormatPattern 99; Unit h
      ProcessValue <- "504_Tank Grouping_DB2020_Time Left Tank_Time Left h Tank 1"
   IOField "I/O field_9" at 128,90 size 42x25; FormatPattern 99; Unit d
      ProcessValue <- "504_Tank Grouping_DB2020_Time Left Tank_Time Left d Tank 1"

PopupScreen "IGG Control from CCR Warning" 665x230
   Button "Button_1" at 0,0 size 665x230; TextOff 'Inert Gas Generator Control Restricted to IGG Room'
      on Click: function_efd93a16("IGG Control from CCR Warning", 0, 0, -1, -1, 1)

screen "Inert Gas Generator Plant" 1280x800, template "Template"
   GraphicView "Graphic view_52" at 522,118 size 43x67; Picture "Graphic_72"
   GraphicView "Graphic view_49" at 715,199 size 43x67; Picture "Graphic_72"
   GraphicView "Graphic view_12" at 522,199 size 43x67; Picture "Graphic_72"
   GraphicView "Graphic view_55" at 522,416 size 43x67; Picture "Graphic_72"
   GraphicView "Graphic view_56" at 650,416 size 43x67; Picture "Graphic_72"
   GraphicView "Graphic view_57" at 522,311 size 43x67; Picture "Graphic_72"
   GraphicView "Graphic view_61" at 527,525 size 32x54; Picture "Graphic_72"
   TextField "Text field_97" at 742,724 size 131x20; Text 'IGG Gas Pressure'
   TextField "Text field_98" at 866,724 size 147x20; Text 'Atom. Air Pressure'
   TextField "Text field_47" at 251,73 size 69x18; Text 'Full Auto'
      Visibility <- "82_To_HMI_CRNT_MODE_IGG"
   TextField "Text field_1" at 251,74 size 55x18; Text 'Manual'
      Visibility <- "82_To_HMI_CRNT_MODE_IGG"
   TextField "Text field_4" at 252,74 size 103x18; Text 'Undetermined'
      Visibility <- "82_To_HMI_CRNT_MODE_IGG"
   TextField "Text field_57" at 252,74 size 36x18; Text 'FAT'
      Visibility <- "82_To_HMI_CRNT_MODE_IGG"
   GraphicView "Logo" at 1,1 size 219x60; Picture "Logo of IGG HMI"
   Group "Group_8" at 743,722 size 397x61
   Button "Button_1" at 902,751 size 66x25; TextOn 'Enabled'; TextOff 'Text'
   IOField "I/O field_29" at 898,751 size 70x25; Authorization "Commissioning"; FormatPattern 99.99; Unit  bar
      ProcessValue <- "1111_PID_CV111_Setpoint"
   Group "Group" at 742,724 size 271x20
   IOField "I/O field_10" at 956,109 size 54x22; FormatPattern 999; Unit %
      ProcessValue <- "12_AI_Data_CV403_SCALED"
   IOField "I/O field_15" at 956,95 size 54x22; FormatPattern 999; Unit %
      ProcessValue <- "16_AQ_Data_CV403_CNTRL"
   GraphicView "Graphic view_5" at 1149,212 size 128x29; Picture "Graphic_82"
   GraphicView "Graphic view_91" at 22,264 size 113x127; Picture "Graphic_246"
   GraphicIOField "Graphic I/O field_5" at 14,257 size 129x139; PictureList "New IA Compressor"
      Visibility <- "68_Sys_Status_Data_IA_PRES_IN_RNG(1)"
      ProcessValue <- "82_To_HMI_IA Compressor Animation"
   GraphicView "Graphic view_93" at 147,261 size 48x132; Picture "Graphic_248"
   TextField "Text field_58" at 41,731 size 135x20; Text 'Fuel Pump System'
      Appearance <- "68_Sys_Status_Data_FUEL_PRES_IN_RNG"
   TextField "Text field_89" at 1115,538 size 54x22; Text 'Text'
   Button "HmiScreenItemData_1" at 1,50 size 150x43; TextOn 'Back'; TextOff 'Main Index'
      on Release: ActivateScreen("02 Main Index", 0)
   GraphicView "Graphic view_20" at 336,126 size 900x542; Picture "IGG_5"
   GraphicView "Graphic view_41" at 815,266 size 13x60; Picture "Graphic_57"
   GraphicView "Graphic view_11" at 296,251 size 377x12; Picture "Graphic_20"
   GraphicView "Graphic view_40" at 806,251 size 21x20; Picture "Graphic_41"
   GraphicView "Graphic view_42" at 296,468 size 278x12; Picture "Graphic_20"
   GraphicView "Graphic view_43" at 696,458 size 19x21; Picture "Graphic_40"
   GraphicView "Graphic view_44" at 294,251 size 20x20; Picture "Graphic_42"
   GraphicView "Graphic view_47" at 295,464 size 11x20; Picture "Graphic_56"
   Group "Group_4" at 522,199 size 43x62; Picture "Graphic_72"
   GraphicView "Graphic view_53" at 313,420 size 43x63; Picture "Graphic_72"
   Group "Group_5" at 522,416 size 43x62; Picture "Graphic_72"
   TextField "Text field_2" at 440,182 size 51x16; Text 'FS-123'
   TextField "Text field_3" at 517,182 size 53x16; Text 'CV-124'
   TextField "Text field_5" at 517,263 size 53x16; Text 'CV-215'
   TextField "Text field_7" at 308,375 size 53x16; Text 'CV-111'
   TextField "Text field_8" at 309,479 size 50x16; Text 'CV-203'
   TextField "Text field_9" at 365,479 size 56x16; Text 'PIT-205'
   TextField "Text field_10" at 518,479 size 50x16; Text 'CV-206'
   TextField "Text field_11" at 646,479 size 50x16; Text 'CV-207'
   TextField "Text field_12" at 364,375 size 59x16; Text 'PIT-113'
   TextField "Text field_13" at 441,375 size 48x16; Text 'FS-115'
   TextField "Text field_14" at 517,375 size 53x16; Text 'CV-114'
   GraphicView "Graphic view_15" at 455,338 size 20x26; Picture "Graphic_79"
   GraphicView "Graphic view_16" at 383,339 size 20x26; Picture "Graphic_36"
   GraphicView "Graphic view_51" at 383,444 size 20x26; Picture "Graphic_36"
   TextField "Text field_21" at 80,649 size 55x18; Text 'E-500B'
   GraphicView "Graphic view_2" at 46,502 size 123x15; Picture "Graphic_99"
   GraphicIOField "Graphic I/O field_3" at 75,482 size 60x65; PictureList "Pump Ani"
      ProcessValue <- "82_To_HMI_Fuel Pump 1 Animation"
   GraphicView "Graphic view_6" at 45,604 size 124x15; Picture "Graphic_99"
   GraphicIOField "Graphic I/O field_4" at 75,585 size 60x65; PictureList "Pump Ani"
      ProcessValue <- "82_To_HMI_Fuel Pump 2 Animation"
   GraphicView "Graphic view_8" at 30,517 size 15x94; Picture "Graphic_101"
   GraphicView "Graphic view_9" at 31,593 size 21x25; Picture "Graphic_96"
   GraphicView "Graphic view_10" at 31,503 size 24x23; Picture "Graphic_102"
   GraphicView "Graphic view_25" at 170,517 size 15x94; Picture "Graphic_101"
   GraphicView "Graphic view_26" at 160,503 size 24x23; Picture "Graphic_104"
   GraphicView "Graphic view_29" at 159,594 size 25x24; Picture "Graphic_97"
   GraphicView "Graphic view_30" at 171,553 size 19x24; Picture "Graphic_103"
   GraphicView "Graphic view_33" at 183,557 size 111x15; Picture "Graphic_99"
   GraphicView "Graphic view_48" at 60,502 size 18x15; Picture "Graphic_99"
   GraphicView "Graphic view_58" at 60,604 size 18x15; Picture "Graphic_99"
   TextField "Text field_22" at 80,549 size 56x18; Text 'E-500A'
   GraphicView "Graphic view_76" at 236,534 size 20x26; Picture "Graphic_36"
   IOField "I/O field_1" at 211,512 size 75x18; FormatPattern s99.99; Unit  Bar
      ProcessValue <- "12_AI_Data_PIT204In_SCALED"
   TextField "Text field_23" at 218,576 size 56x16; Text 'PIT-204'
   Rectangle "Rectangle_9" at 66,477 size 78x92
      Appearance <- "10_DI_Data_E500A_TRIPPED"
   Rectangle "Rectangle_10" at 66,580 size 79x92
      Appearance <- "10_DI_Data_E500B_TRIPPED(1)"
   TextField "Text field_24" at 67,673 size 83x18; Text 'Duty Pump'
      Visibility <- "101_Fuel_Pumps_DB_Duty Is B"
   TextField "Text field_25" at 67,457 size 83x18; Text 'Duty Pump'
      Visibility <- "101_Fuel_Pumps_DB_Duty Is A"
   Circle "Circle_11" at 35,559 size 6x6
      Visibility <- "10_DI_Data_E500A_ENBLD"
   GraphicView "Graphic view_46" at 285,547 size 20x24; Picture "Graphic_40"
   GraphicView "Graphic view_21" at 789,331 size 24x10; Picture "Graphic_63"
   GraphicView "Graphic view_22" at 785,326 size 12x13; Picture "Graphic_64"
   GraphicView "Graphic view_23" at 784,176 size 9x156; Picture "Graphic_70"
   GraphicView "Graphic view_27" at 279,176 size 9x185; Picture "Graphic_70"
   GraphicView "Graphic view_35" at 281,363 size 325x11; Picture "Graphic_63"
   GraphicView "Graphic view_39" at 687,379 size 8x10; Picture "Graphic_70"
   GraphicView "Graphic view_38" at 688,386 size 10x13; Picture "Graphic_64"
   GraphicView "Graphic view_7" at 455,147 size 20x26; Picture "Graphic_79"
   GraphicView "Graphic view_18" at 780,172 size 13x15; Picture "Graphic_67"
   GraphicView "Graphic view_14" at 281,171 size 318x11; Picture "Graphic_63"
   GraphicView "Graphic view_17" at 279,172 size 13x15; Picture "Graphic_66"
   Group "Group_2" at 522,118 size 43x62; Picture "Graphic_72"
   GraphicView "Graphic view_31" at 236,331 size 20x26; Picture "Graphic_36"
   IOField "I/O field_6" at 207,308 size 74x18; FormatPattern s99.99; Unit  Bar
      ProcessValue <- "12_AI_Data_PIT112In_SCALED"
   TextField "Text field_17" at 218,375 size 56x16; Text 'PIT-112'
   GraphicView "Graphic view_50" at 313,314 size 43x63; Picture "Graphic_72"
   Group "Group_7" at 522,311 size 43x62; Picture "Graphic_72"
   GraphicView "Graphic view_45" at 293,262 size 13x297; Picture "Graphic_57"
   GraphicView "Graphic view_54" at 305,517 size 24x21; Picture "Graphic_107"
   IOField "I/O field_7" at 358,423 size 77x18; FormatPattern s99.99; Unit  bar
      ProcessValue <- "12_AI_Data_PIT205In_SCALED"
   TextField "Text field_18" at 513,418 size 60x22; Text 'Closed'
      Visibility <- "14_DQ_Data_200CV206ControlOut"
   TextField "Text field_19" at 513,418 size 60x22; Text 'Opened'
      Visibility <- "14_DQ_Data_200CV206ControlOut"
   IOField "I/O field_11" at 330,522 size 55x18; FormatPattern 99.9; Unit  °C
      ProcessValue <- "12_AI_Data_TIT202In_SCALED"
   GraphicView "Graphic view_59" at 558,468 size 145x12; Picture "Graphic_20"
   TextField "Text field_20" at 514,200 size 60x22; Text 'Closed'
   TextField "Text field_26" at 514,200 size 60x22; Text 'Opened'
      Visibility <- "14_DQ_Data_200CV215ControlOut"
   TextField "Text field_31" at 513,315 size 60x22; Text 'Closed'
   TextField "Text field_32" at 513,315 size 60x22; Text 'Opened'
      Visibility <- "14_DQ_Data_200CV114ControlOut"
   TextField "Text field_33" at 305,541 size 56x16; Text 'TIT-202'
   GraphicView "Graphic view_62" at 647,251 size 173x12; Picture "Graphic_20"
   Group "Group_6" at 650,416 size 43x62; Picture "Graphic_72"
   GraphicView "Graphic view_34" at 705,425 size 11x43; Picture "Graphic_57"
   TextField "Text field_28" at 641,419 size 60x22; Text 'Closed'
   TextField "Text field_29" at 641,419 size 60x22; Text 'Opened'
      Visibility <- "14_DQ_Data_200CV207ControlOut"
   GraphicView "Graphic view_63" at 565,171 size 223x11; Picture "Graphic_63"
   Group "Group_3" at 715,199 size 43x62; Picture "Graphic_72"
   TextField "Text field_6" at 710,263 size 53x16; Text 'CV-216'
   TextField "Text field_27" at 706,200 size 60x22; Text 'Closed'
   TextField "Text field_30" at 706,200 size 60x22; Text 'Opened'